REGION Network 32: "MFC-4024-T_DB"
   RUNG wire#powerrail
      "MFC-4024-T_DB"(Mode := 2, RAIVI :=, RAIVR :=, EnableHighAlarms :=, EnableLowAlarms :=, "TI Fail" :=, SAI =>)
   END_RUNG
   RUNG wire#powerrail
      I_Contact( false )
      { S7_GenerateENO := "TRUE" } Move(in := "MFC-4024_MB_R_DB".MB_Data.Buffer[2], out1 => "MFC-4024-T_DB".RAIVR)
   END_RUNG
   // the same network as SCL:
   "MFC-4024-T_DB"(Mode := 2);   // "TX-AI"
   IF NOT false THEN "MFC-4024-T_DB".RAIVR := "MFC-4024_MB_R_DB".MB_Data.Buffer[2]; END_IF;
END_REGION

REGION Network 33: "MFC-4025-T_DB"
   RUNG wire#powerrail
      "MFC-4025-T_DB"(Mode := 2, RAIVI :=, RAIVR :=, EnableHighAlarms :=, EnableLowAlarms :=, "TI Fail" :=, SAI =>)
   END_RUNG
   RUNG wire#powerrail
      I_Contact( false )
      { S7_GenerateENO := "TRUE" } Move(in := "MFC-4025_MB_R_DB".MB_Data.Buffer[2], out1 => "MFC-4025-T_DB".RAIVR)
   END_RUNG
   // the same network as SCL:
   "MFC-4025-T_DB"(Mode := 2);   // "TX-AI"
   IF NOT false THEN "MFC-4025-T_DB".RAIVR := "MFC-4025_MB_R_DB".MB_Data.Buffer[2]; END_IF;
END_REGION
END_FUNCTION

// folder: Analogs inputs/Trasmitters/VFD_Feedback Trasmitters

FUNCTION "VFDFeedbackTrasmitters" : Void   // FC14, LAD
TITLE = VFD Feedback
{ S7_Optimized_Access := 'TRUE' }
VERSION : 0.1
// Updated Date:
// Note:
   VAR_TEMP
      Alarms : Struct
         "T-101_AlarmsEnab" : Bool;
         "T-102_AlarmsEnab" : Bool;
         "R-201_AlarmsEnab" : Bool;
         "R-202_AlarmsEnab" : Bool;
         Centrifuge_AlarmsEnab : Bool;
      END_STRUCT;
      temporalvar : Int;
   END_VAR
BEGIN

REGION Network 1: Enable T-101 Agitator Alarms
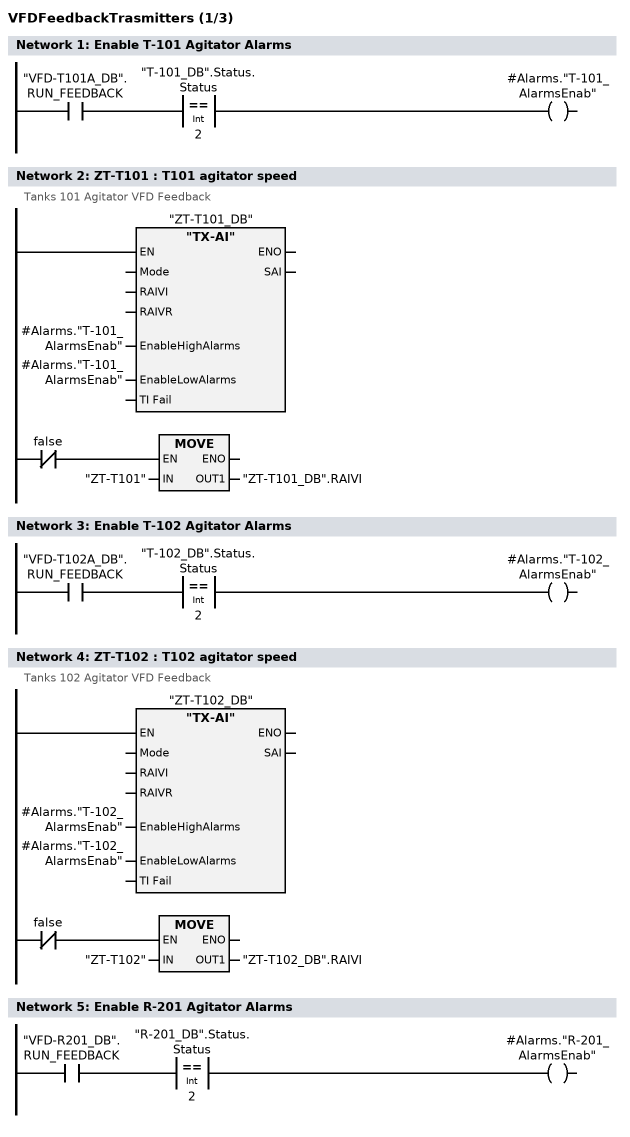
   RUNG wire#powerrail
      Contact( "VFD-T101A_DB".RUN_FEEDBACK )
      { S7_Templates := "SrcType := Int" } EQ_Contact(in1 := "T-101_DB".Status.Status, in2 := 2)
      Coil( #Alarms."T-101_AlarmsEnab" )
   END_RUNG
   // the same network as SCL:
   #Alarms."T-101_AlarmsEnab" := "VFD-T101A_DB".RUN_FEEDBACK AND ("T-101_DB".Status.Status = 2);
END_REGION

REGION Network 2: ZT-T101 : T101 agitator speed
   // Tanks 101 Agitator VFD Feedback
   RUNG wire#powerrail
      "ZT-T101_DB"(Mode :=, RAIVI :=, RAIVR :=, EnableHighAlarms := #Alarms."T-101_AlarmsEnab", EnableLowAlarms := #Alarms."T-101_AlarmsEnab", "TI Fail" :=, SAI =>)
   END_RUNG
   RUNG wire#powerrail
      I_Contact( false )
      { S7_GenerateENO := "TRUE" } Move(in := "ZT-T101", out1 => "ZT-T101_DB".RAIVI)
   END_RUNG
   // the same network as SCL:
   "ZT-T101_DB"(EnableHighAlarms := #Alarms."T-101_AlarmsEnab", EnableLowAlarms := #Alarms."T-101_AlarmsEnab");   // "TX-AI"
   IF NOT false THEN "ZT-T101_DB".RAIVI := "ZT-T101"; END_IF;
END_REGION

REGION Network 3: Enable T-102 Agitator Alarms
   RUNG wire#powerrail
      Contact( "VFD-T102A_DB".RUN_FEEDBACK )
      { S7_Templates := "SrcType := Int" } EQ_Contact(in1 := "T-102_DB".Status.Status, in2 := 2)
      Coil( #Alarms."T-102_AlarmsEnab" )
   END_RUNG
   // the same network as SCL:
   #Alarms."T-102_AlarmsEnab" := "VFD-T102A_DB".RUN_FEEDBACK AND ("T-102_DB".Status.Status = 2);
END_REGION

REGION Network 4: ZT-T102 : T102 agitator speed
   // Tanks 102 Agitator VFD Feedback
   RUNG wire#powerrail
      "ZT-T102_DB"(Mode :=, RAIVI :=, RAIVR :=, EnableHighAlarms := #Alarms."T-102_AlarmsEnab", EnableLowAlarms := #Alarms."T-102_AlarmsEnab", "TI Fail" :=, SAI =>)
   END_RUNG
   RUNG wire#powerrail
      I_Contact( false )
      { S7_GenerateENO := "TRUE" } Move(in := "ZT-T102", out1 => "ZT-T102_DB".RAIVI)
   END_RUNG
   // the same network as SCL:
   "ZT-T102_DB"(EnableHighAlarms := #Alarms."T-102_AlarmsEnab", EnableLowAlarms := #Alarms."T-102_AlarmsEnab");   // "TX-AI"
   IF NOT false THEN "ZT-T102_DB".RAIVI := "ZT-T102"; END_IF;
END_REGION

REGION Network 5: Enable R-201 Agitator Alarms
   RUNG wire#powerrail
      Contact( "VFD-R201_DB".RUN_FEEDBACK )
      { S7_Templates := "SrcType := Int" } EQ_Contact(in1 := "R-201_DB".Status.Status, in2 := 2)
      Coil( #Alarms."R-201_AlarmsEnab" )
   END_RUNG
   // the same network as SCL:
   #Alarms."R-201_AlarmsEnab" := "VFD-R201_DB".RUN_FEEDBACK AND ("R-201_DB".Status.Status = 2);
END_REGION

REGION Network 6: ZT-R201 : R201 agitator speed
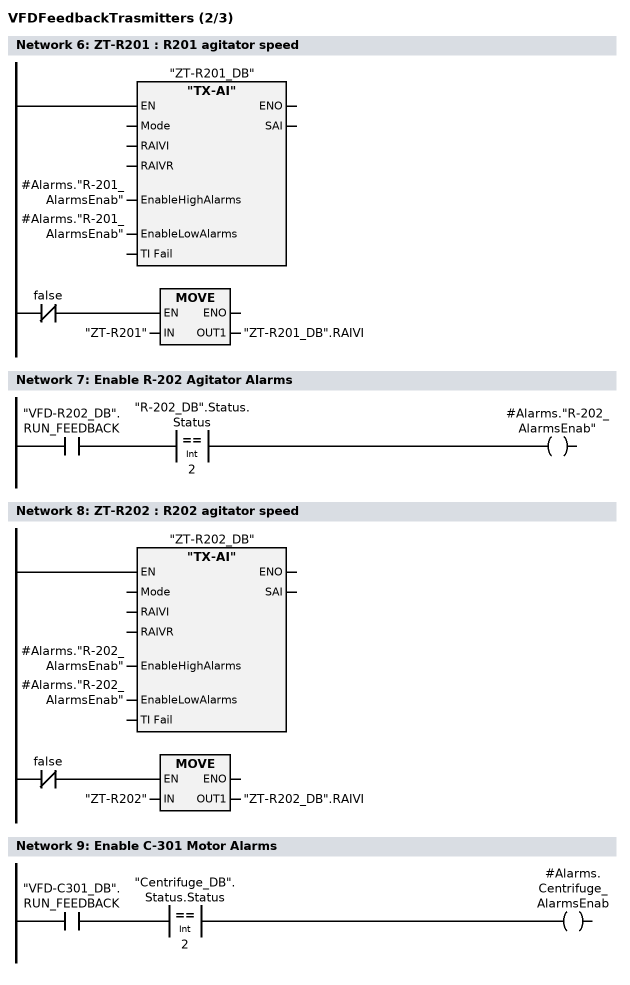
   RUNG wire#powerrail
      "ZT-R201_DB"(Mode :=, RAIVI :=, RAIVR :=, EnableHighAlarms := #Alarms."R-201_AlarmsEnab", EnableLowAlarms := #Alarms."R-201_AlarmsEnab", "TI Fail" :=, SAI =>)
   END_RUNG
   RUNG wire#powerrail
      I_Contact( false )
      { S7_GenerateENO := "TRUE" } Move(in := "ZT-R201", out1 => "ZT-R201_DB".RAIVI)
   END_RUNG
   // the same network as SCL:
   "ZT-R201_DB"(EnableHighAlarms := #Alarms."R-201_AlarmsEnab", EnableLowAlarms := #Alarms."R-201_AlarmsEnab");   // "TX-AI"
   IF NOT false THEN "ZT-R201_DB".RAIVI := "ZT-R201"; END_IF;
END_REGION

REGION Network 7: Enable R-202 Agitator Alarms
   RUNG wire#powerrail
      Contact( "VFD-R202_DB".RUN_FEEDBACK )
      { S7_Templates := "SrcType := Int" } EQ_Contact(in1 := "R-202_DB".Status.Status, in2 := 2)
      Coil( #Alarms."R-202_AlarmsEnab" )
   END_RUNG
   // the same network as SCL:
   #Alarms."R-202_AlarmsEnab" := "VFD-R202_DB".RUN_FEEDBACK AND ("R-202_DB".Status.Status = 2);
END_REGION

REGION Network 8: ZT-R202 : R202 agitator speed
   RUNG wire#powerrail
      "ZT-R202_DB"(Mode :=, RAIVI :=, RAIVR :=, EnableHighAlarms := #Alarms."R-202_AlarmsEnab", EnableLowAlarms := #Alarms."R-202_AlarmsEnab", "TI Fail" :=, SAI =>)
   END_RUNG
   RUNG wire#powerrail
      I_Contact( false )
      { S7_GenerateENO := "TRUE" } Move(in := "ZT-R202", out1 => "ZT-R202_DB".RAIVI)
   END_RUNG
   // the same network as SCL:
   "ZT-R202_DB"(EnableHighAlarms := #Alarms."R-202_AlarmsEnab", EnableLowAlarms := #Alarms."R-202_AlarmsEnab");   // "TX-AI"
   IF NOT false THEN "ZT-R202_DB".RAIVI := "ZT-R202"; END_IF;
END_REGION

REGION Network 9: Enable C-301 Motor Alarms
   RUNG wire#powerrail
      Contact( "VFD-C301_DB".RUN_FEEDBACK )
      { S7_Templates := "SrcType := Int" } EQ_Contact(in1 := "Centrifuge_DB".Status.Status, in2 := 2)
      Coil( #Alarms.Centrifuge_AlarmsEnab )
   END_RUNG
   // the same network as SCL:
   #Alarms.Centrifuge_AlarmsEnab := "VFD-C301_DB".RUN_FEEDBACK AND ("Centrifuge_DB".Status.Status = 2);
END_REGION

REGION Network 10: ZT-C-301 : C-301 Motorspeed
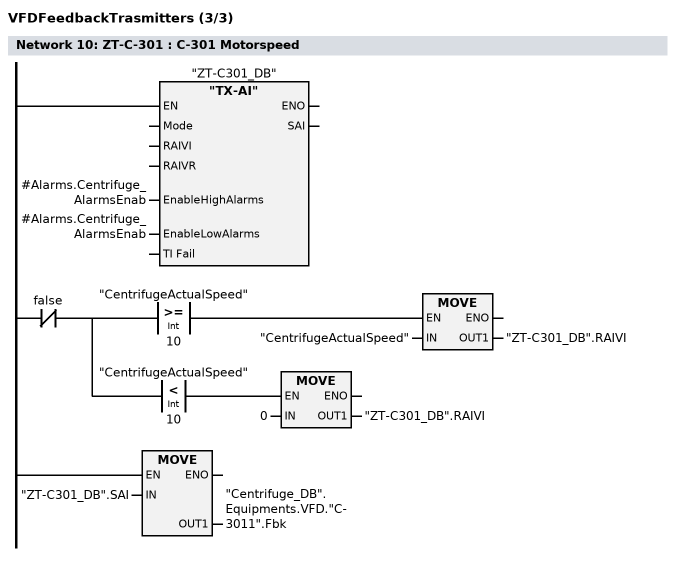
   RUNG wire#powerrail
      "ZT-C301_DB"(Mode :=, RAIVI :=, RAIVR :=, EnableHighAlarms := #Alarms.Centrifuge_AlarmsEnab, EnableLowAlarms := #Alarms.Centrifuge_AlarmsEnab, "TI Fail" :=, SAI =>)
   END_RUNG
   RUNG wire#powerrail
      I_Contact( false )
      wire#w1
      { S7_Templates := "SrcType := Int" } GE_Contact(in1 := "CentrifugeActualSpeed", in2 := 10)
      { S7_GenerateENO := "TRUE" } Move(in := "CentrifugeActualSpeed", out1 => "ZT-C301_DB".RAIVI)
   END_RUNG
   RUNG wire#w1
      { S7_Templates := "SrcType := Int" } LT_Contact(in1 := "CentrifugeActualSpeed", in2 := 10)
      { S7_GenerateENO := "TRUE" } Move(in := 0, out1 => "ZT-C301_DB".RAIVI)
   END_RUNG
   RUNG wire#powerrail
      Move(in := "ZT-C301_DB".SAI, out1 => "Centrifuge_DB".Equipments.VFD."C-3011".Fbk)
   END_RUNG
   // the same network as SCL:
   "ZT-C301_DB"(EnableHighAlarms := #Alarms.Centrifuge_AlarmsEnab,   // "TX-AI"
                EnableLowAlarms := #Alarms.Centrifuge_AlarmsEnab);
   IF NOT false AND ("CentrifugeActualSpeed" >= 10) THEN
       "ZT-C301_DB".RAIVI := "CentrifugeActualSpeed";
   END_IF;
   IF NOT false AND ("CentrifugeActualSpeed" < 10) THEN "ZT-C301_DB".RAIVI := 0; END_IF;
   "Centrifuge_DB".Equipments.VFD."C-3011".Fbk := "ZT-C301_DB".SAI;
END_REGION
END_FUNCTION

// folder: Analogs inputs/Trasmitters/Vibration Transmitter

FUNCTION "VibrationTransmitter" : Void   // FC107, LAD
{ S7_Optimized_Access := 'TRUE' }
VERSION : 0.1
BEGIN

REGION Network 1: Centrifuge Vibration Transmitter
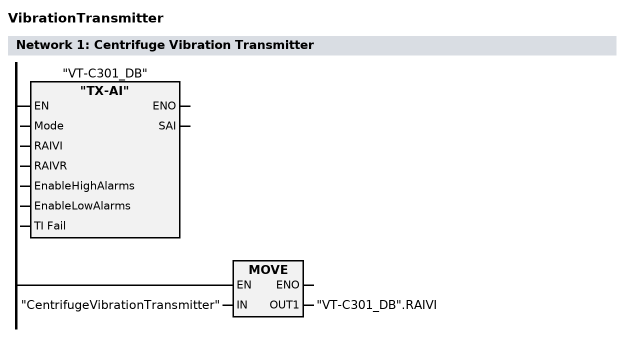
   RUNG wire#powerrail
      "VT-C301_DB"(Mode :=, RAIVI :=, RAIVR :=, EnableHighAlarms :=, EnableLowAlarms :=, "TI Fail" :=, SAI =>)
   END_RUNG
   RUNG wire#powerrail
      Move(in := "CentrifugeVibrationTransmitter", out1 => "VT-C301_DB".RAIVI)
   END_RUNG
   // the same network as SCL:
   "VT-C301_DB"();   // "TX-AI"
   "VT-C301_DB".RAIVI := "CentrifugeVibrationTransmitter";
END_REGION
END_FUNCTION

// folder: Calculations

FUNCTION_BLOCK "Array_Intergration"   // FB21, LAD
TITLE = Level to VFD Table
{ S7_Optimized_Access := 'TRUE' }
VERSION : 0.1
// Level to V FD Interpolation Table
   VAR_INPUT
      PV : Real;
      Ramp_UP : Bool := True;   // Ramp Up Sequence Enable
      Ramp_Down : Bool;   // Ramp Down Sequence Enable
   END_VAR
   VAR_OUTPUT
      SP : Real;
   END_VAR
   VAR
      FirstScan : Bool := TRUE;
      Number : UInt;
      "Array" : Array[0..#Array_Size] of Struct
         X : Real;   // Set Point for Level
         Y : Real;   // Output to Drive VFD
         X1 : Real;
         X2 : Real;
         Y1 : Real;
      END_STRUCT;
      TP_Up : IEC_TIMER;
      TP_Down : IEC_TIMER;
      Deadband : Struct
         UDW : Real := 0.5;   // Upper Deadband Width
         LDW : Real := 0.5;   // Lower Deadband Width
      END_STRUCT;
   END_VAR
   VAR_TEMP
      Trigger : Array[0..1] of Bool;
      Deadband_SP : Struct
         UDW : Real;   // Upper Deadband Width
         LDW : Real;   // Lower Deadband Width
      END_STRUCT;
      temp_CAl : Array[0..#Temp_Count] of Real;
   END_VAR
   VAR CONSTANT
      Array_Size : UInt := 4;
      TRigger_Count : UInt := 2;
      Temp_Count : UInt := 4;
   END_VAR
   VAR_TEMP   // added for the SCL form of the ladder/FBD networks
      _w1 : Bool;
      _w2 : Bool;
   END_VAR
   // "Array"[1].X := 20.0;
   // "Array"[2].X := 30.0;
   // "Array"[3].X := 40.0;
   // "Array"[4].X := 50.0;
   // TP_Up.PT := T#1ms;
   // TP_Down.PT := T#500ms;
BEGIN

REGION Network 1: First Scan
   // First Scan  Set array to Begining of the Table
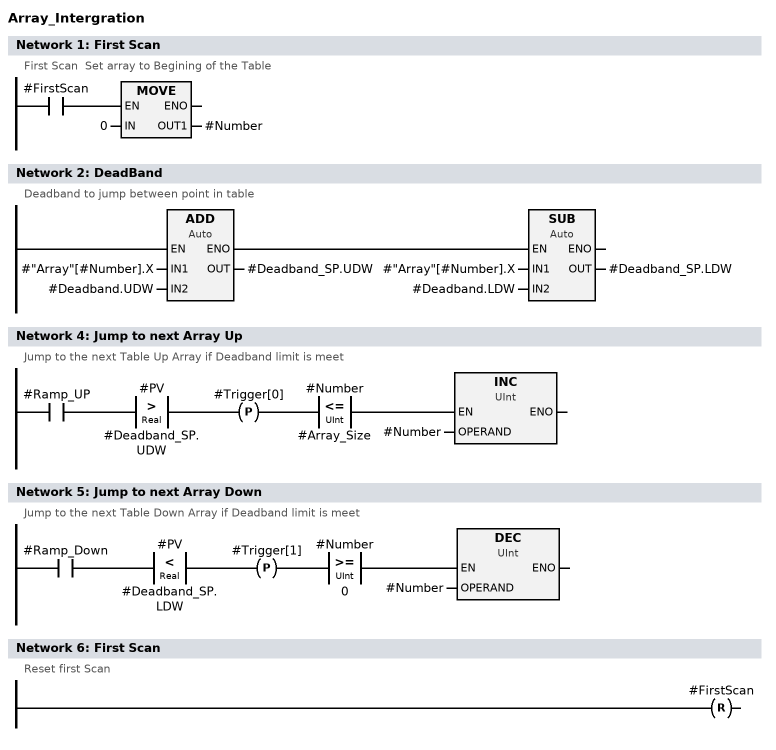
   RUNG wire#powerrail
      Contact( #FirstScan )
      { S7_GenerateENO := "TRUE" } Move(in := 0, out1 => #Number)
   END_RUNG
   // the same network as SCL:
   IF #FirstScan THEN #Number := 0; END_IF;
END_REGION

REGION Network 2: DeadBand
   // Deadband to jump between point in table
   RUNG wire#powerrail
      { S7_GenerateENO := "TRUE" } Add(in1 := #"Array"[#Number].X, in2 := #Deadband.UDW, out => #Deadband_SP.UDW)
      { S7_GenerateENO := "TRUE" } Sub(in1 := #"Array"[#Number].X, in2 := #Deadband.LDW, out => #Deadband_SP.LDW)
   END_RUNG
   // the same network as SCL:
   // ENO of a box is taken as its EN; it also drops when the box reports an error
   #Deadband_SP.UDW := #"Array"[#Number].X + #Deadband.UDW;
   #Deadband_SP.LDW := #"Array"[#Number].X - #Deadband.LDW;
END_REGION

REGION Network 3 (SCL): Table Calculation
   // Interpolation Formula implementation if the Ramp sequence is on and Deadband
   IF #Ramp_UP=TRUE AND #PV<=#Deadband_SP.UDW THEN
       // Interpolation Formula
       // Y = Y1 + (Y2 – Y1)/(X2 – X1) * (X * X1)
       #temp_CAl[0] := #Array[#Number].X * #Array[#Number].X1;// (X * X1)
       #temp_CAl[1] := #Array[#Number].X2 * #Array[#Number].X1;// (X2 – X1)
       #temp_CAl[2] := #Array[#Number].X2 * #Array[#Number].X1;// (Y2 – Y1)
       #temp_CAl[3] := #temp_CAl[1] / #temp_CAl[2];//(Y2 – Y1)/(X2 – X1)
       #temp_CAl[4] := #temp_CAl[3] * #temp_CAl[0];
       #SP := #Array[#Number].Y1 + #temp_CAl[4]; //SUM
   END_IF;
   IF #Ramp_Down=TRUE AND #PV>=#Deadband_SP.LDW THEN
       // Interpolation Formula
       // Y = Y1 + (Y2 – Y1)/(X2 – X1) * (X * X1)
       #temp_CAl[0] := #Array[#Number].X * #Array[#Number].X1;// (X * X1)
       #temp_CAl[1] := #Array[#Number].X2 * #Array[#Number].X1;// (X2 – X1)
       #temp_CAl[2] := #Array[#Number].X2 * #Array[#Number].X1;// (Y2 – Y1)
       #temp_CAl[3] := #temp_CAl[1] / #temp_CAl[2];//(Y2 – Y1)/(X2 – X1)
       #temp_CAl[4] := #temp_CAl[3] * #temp_CAl[0];
       #SP := #Array[#Number].Y1 + #temp_CAl[4]; //SUM
   END_IF;
END_REGION

REGION Network 4: Jump to next Array Up
   // Jump to the next Table Up Array if Deadband limit is meet
   RUNG wire#powerrail
      Contact( #Ramp_UP )
      { S7_Templates := "SrcType := Real" } GT_Contact(in1 := #PV, in2 := #Deadband_SP.UDW)
      P_Trig( #Trigger[0] )
      { S7_Templates := "SrcType := UInt" } LE_Contact(in1 := #Number, in2 := #Array_Size)
      { S7_Templates := "DestType := UInt"; S7_GenerateENO := "TRUE" } Inc( #Number )
   END_RUNG
   // the same network as SCL:
   #_w1 := #Ramp_UP AND (#PV > #Deadband_SP.UDW);
   #_w2 := #_w1 AND NOT #Trigger[0];   // rising edge
   #Trigger[0] := #_w1;
   IF #_w2 AND (#Number <= #Array_Size) THEN #Number := #Number + 1; END_IF;
END_REGION

REGION Network 5: Jump to next Array Down
   // Jump to the next Table Down Array if Deadband limit is meet
   RUNG wire#powerrail
      Contact( #Ramp_Down )
      { S7_Templates := "SrcType := Real" } LT_Contact(in1 := #PV, in2 := #Deadband_SP.LDW)
      P_Trig( #Trigger[1] )
      { S7_Templates := "SrcType := UInt" } GE_Contact(in1 := #Number, in2 := 0)
      { S7_Templates := "DestType := UInt"; S7_GenerateENO := "TRUE" } Dec( #Number )
   END_RUNG
   // the same network as SCL:
   #_w1 := #Ramp_Down AND (#PV < #Deadband_SP.LDW);
   #_w2 := #_w1 AND NOT #Trigger[1];   // rising edge
   #Trigger[1] := #_w1;
   IF #_w2 AND (#Number >= 0) THEN #Number := #Number - 1; END_IF;
END_REGION

REGION Network 6: First Scan
   // Reset first Scan
   RUNG wire#powerrail
      R_Coil( #FirstScan )
   END_RUNG
   // the same network as SCL:
   #FirstScan := FALSE;
END_REGION
END_FUNCTION_BLOCK

FUNCTION_BLOCK "Tank_Calculation_FB"   // FB22, LAD
{ S7_Optimized_Access := 'TRUE' }
VERSION : 0.1
   VAR_INPUT
      Mode : UInt;   // Type of Tank mode: 1= Vertical Capsule Tank
      Level : Real;
   END_VAR
   VAR_OUTPUT
      ScaleVolume : Real;
   END_VAR
   VAR
      "Vertical Capsule Tank" : Struct
         Enable : Bool;
         "case" : USInt;   // Mode: | Vcylpartial=1 | Vcylpartial & Vbottom_head_partial = 2 | Vcylpartial & Vtop_head_partial = 3 | Vcyl_total = 4 |
         Static_1 : USInt;   // tank internal diameter
         DiameterCylindrical : UInt;
         Height : UInt;
      END_STRUCT;
   END_VAR
   VAR_TEMP
      "Case" : USInt;
      Vcylpartial : Real;
      TEmp : Real;
      temp_CAl : Array[0..#Temp_Count] of Real;
   END_VAR
   VAR CONSTANT
      "Vertical Capsule Tank_1" : UInt := 1;
      MAthPi : Real := 3.14;
      Temp_Count : UInt := 4;
   END_VAR
BEGIN

REGION Network 1: Mode1: Selected
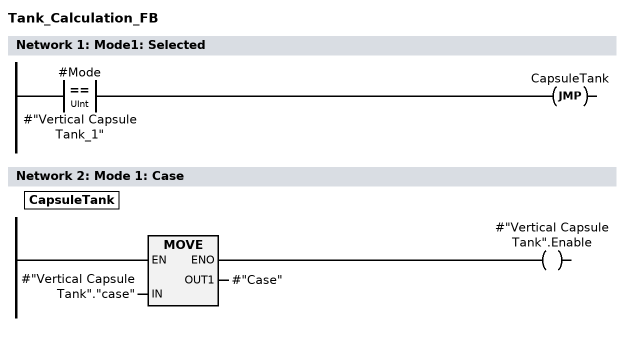
   RUNG wire#powerrail
      { S7_Templates := "SrcType := UInt" } EQ_Contact(in1 := #Mode, in2 := #"Vertical Capsule Tank_1")
      JumpCoil( CapsuleTank )
   END_RUNG
   // the same network as SCL:
   IF #Mode = #"Vertical Capsule Tank_1" THEN GOTO CapsuleTank; END_IF;
END_REGION

REGION Network 2: Mode 1: Case
   Label( CapsuleTank )
   RUNG wire#powerrail
      { S7_GenerateENO := "TRUE" } Move(in := #"Vertical Capsule Tank"."case", out1 => #"Case")
      Coil( #"Vertical Capsule Tank".Enable )
   END_RUNG
   // the same network as SCL:
   // ENO of a box is taken as its EN; it also drops when the box reports an error
   CapsuleTank:
   #"Case" := #"Vertical Capsule Tank"."case";
   #"Vertical Capsule Tank".Enable := TRUE;
END_REGION

REGION Network 3 (SCL): Vertical Capsule Tank CAlculation
   CASE #Case OF
       1:(*Mode:Partial Volume horizontal Cylinderical Calculation
       Note: Calculation For the cylindrical part Of the tank only 
             does not Contain Top Head or Botton Head of vessel
       Formula: Vcylpartial=π*〖ID〗^2/4*Lv*)
           #temp_CAl[0] := #"Vertical Capsule Tank".DiameterCylindrical / 2;//Radius /cylindrical
           #temp_CAl[1] := #MAthPi * #temp_CAl[0] ** 2 * (#Level - 2 * #temp_CAl[0]);// Volume Cylinderical  
           #temp_CAl[2] := #Level/ (#MAthPi * #temp_CAl[0] ** 2);// Liquid Level
           #Vcylpartial := #Level - (#temp_CAl[2]);// Current Level
           #ScaleVolume := #Vcylpartial;// Move To Volume
           ;
       2:  (*Mode: The liquid level is in the Botton head of the vessel to the top of the Cylinderical part of the Vessel the top head of the Vessel not  *)
           IF #Level >= 0 AND #Level <= 20 THEN
               // From 0 to 20 The liquid level is low, within the bottom head of the vessel
             //  #temp_CAl[0] := #MAthPi/6*(3*)  ;
             //  #Vbottom_head = 
               ;
           ELSE

               ;
           END_IF;


           ;
       3:  // The liquid level is reaching the top head of the vessel
           ;
       ELSE  // Set Case Value to 0
           #Case := 0;
           ;
   END_CASE;
END_REGION
END_FUNCTION_BLOCK

FUNCTION_BLOCK "Array_Intergration_B"   // FB23, LAD
TITLE = Level to VFD Table
{ S7_Optimized_Access := 'TRUE' }
VERSION : 0.1
// Level to V FD Interpolation Table
   VAR_INPUT
      PV : Int;
      Ramp_UP : Bool := True;   // Ramp Up Sequence Enable
      Ramp_Down : Bool;   // Ramp Down Sequence Enable
   END_VAR
   VAR_OUTPUT
      SP : Real;
   END_VAR
   VAR
      FirstScan : Bool := TRUE;
      Number : UInt;
      "X Axis Max" : Int := 100;
      "Y Axis max" : Int := 4000;
      "array of X" : Array[0..#Array_Size] of Int;   // Level Setpoints
      "array of Y" : Array[0..#Array_Size] of Int;   // RPM Sepoints
      "Array" : Array[0..#Array_Size] of Struct
         X : Int;   // Set Point for Level
         Y : Int;   // Output to Drive VFD
         X1 : Int;
         X2 : Int;
         Y1 : Int;
         Y2 : Int;
      END_STRUCT;
      Formula : Struct
         X : Int;   // Set Point for Level
         Y : Int;   // Output to Drive VFD
         X1 : Int;
         X2 : Int;
         Y1 : Int;
         Y2 : Int;
      END_STRUCT;
      TP_Up : IEC_TIMER;
      TP_Down : IEC_TIMER;
      Deadband : Struct
         UDW : Real := 0.5;   // Upper Deadband Width
         LDW : Real := 0.5;   // Lower Deadband Width
      END_STRUCT;
   END_VAR
   VAR_TEMP
      Trigger : Array[0..1] of Bool;
      Deadband_SP : Struct
         UDW : Real;   // Upper Deadband Width
         LDW : Real;   // Lower Deadband Width
      END_STRUCT;
      temp_CAl : Array[0..#Temp_Count] of Real;
   END_VAR
   VAR CONSTANT
      Array_Size : UInt := 4;
      TRigger_Count : UInt := 2;
      Temp_Count : UInt := 5;
      RMP : UInt := 3000;
   END_VAR
   // TP_Up.PT := T#1ms;
   // TP_Down.PT := T#500ms;
   // "array of X"[0] := 20;
   // "array of X"[1] := 30;
   // "array of X"[2] := 40;
   // "array of X"[3] := 50;
   // "array of X"[4] := 60;
   // "array of Y"[0] := 500;
   // "array of Y"[1] := 1000;
   // "array of Y"[2] := 1500;
   // "array of Y"[3] := 2000;
   // "array of Y"[4] := 1500;
BEGIN

REGION Network 1: First Scan
   // First Scan  Set array to Begining of the Table
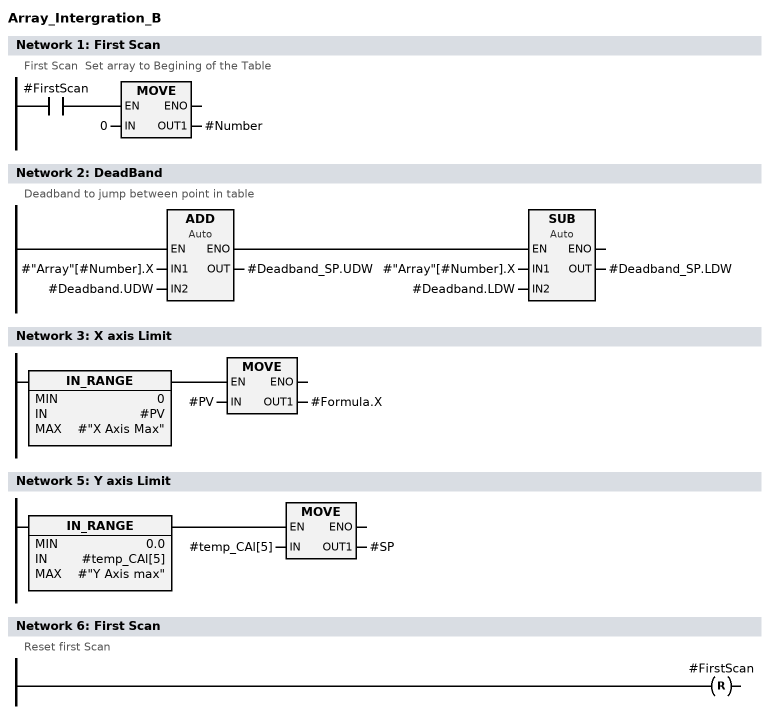
   RUNG wire#powerrail
      Contact( #FirstScan )
      { S7_GenerateENO := "TRUE" } Move(in := 0, out1 => #Number)
   END_RUNG
   // the same network as SCL:
   IF #FirstScan THEN #Number := 0; END_IF;
END_REGION

REGION Network 2: DeadBand
   // Deadband to jump between point in table
   RUNG wire#powerrail
      { S7_GenerateENO := "TRUE" } Add(in1 := #"Array"[#Number].X, in2 := #Deadband.UDW, out => #Deadband_SP.UDW)
      { S7_GenerateENO := "TRUE" } Sub(in1 := #"Array"[#Number].X, in2 := #Deadband.LDW, out => #Deadband_SP.LDW)
   END_RUNG
   // the same network as SCL:
   // ENO of a box is taken as its EN; it also drops when the box reports an error
   #Deadband_SP.UDW := #"Array"[#Number].X + #Deadband.UDW;
   #Deadband_SP.LDW := #"Array"[#Number].X - #Deadband.LDW;
END_REGION

REGION Network 3: X axis Limit
   RUNG wire#powerrail
      { S7_Templates := "SrcType := Int" } InRange(min := 0, in := #PV, max := #"X Axis Max")
      { S7_GenerateENO := "TRUE" } Move(in := #PV, out1 => #Formula.X)
   END_RUNG
   // the same network as SCL:
   IF (0 <= #PV) AND (#PV <= #"X Axis Max") THEN #Formula.X := #PV; END_IF;
END_REGION

REGION Network 4 (SCL): Table Calculation
   // Interpolation Formula implementation if the Ramp sequence is on and Deadband
   // Interpolation Formula
   // Y = Y1 + (Y2 – Y1)/(X2 – X1) * (X * X1)
   #Formula.Y1 := #"array of Y"[0];
   #Formula.X1 := #"array of X"[0];
   #Formula.Y2 := #"array of Y"[1];
   #Formula.X2 := #"array of X"[1];
   #temp_CAl[0] := #Formula.Y2 * #Formula.Y1;// (Y2 – Y1)
   #temp_CAl[1] := #Formula.X2 - #Formula.X1;// (X2 – X1)
   #temp_CAl[2] := #Formula.X * #Formula.X1;// (X * X1)
   #temp_CAl[3] := #temp_CAl[0] / #temp_CAl[1];//(Y2 – Y1)/(X2 – X1)
   #temp_CAl[4] := #temp_CAl[3] * #temp_CAl[2];//(Y2 – Y1)/(X2 – X1) * (X * X1)
   #temp_CAl[5] := #Formula.Y1 + #temp_CAl[4];//Y1 + (Y2 – Y1)/(X2 – X1) * (X * X1)
END_REGION

REGION Network 5: Y axis Limit
   RUNG wire#powerrail
      { S7_Templates := "SrcType := Real" } InRange(min := 0.0, in := #temp_CAl[5], max := #"Y Axis max")
      { S7_GenerateENO := "TRUE" } Move(in := #temp_CAl[5], out1 => #SP)
   END_RUNG
   // the same network as SCL:
   IF (0.0 <= #temp_CAl[5]) AND (#temp_CAl[5] <= #"Y Axis max") THEN #SP := #temp_CAl[5]; END_IF;
END_REGION

REGION Network 6: First Scan
   // Reset first Scan
   RUNG wire#powerrail
      R_Coil( #FirstScan )
   END_RUNG
   // the same network as SCL:
   #FirstScan := FALSE;
END_REGION
END_FUNCTION_BLOCK

FUNCTION_BLOCK "Volume_Calculation"   // FB25, SCL
{ S7_Optimized_Access := 'TRUE' }
VERSION : 0.1
   VAR_INPUT
      Input : Int;
      Input_Max : Real;
      Input_Min : Real;
   END_VAR
   VAR_OUTPUT
      "Volume (L)" : Real;   // Valume in Gallons
      "Volume (Gal)" : Real;   // Volume in Liters
   END_VAR
   VAR
      CurrentCylinderVolume : Struct   // Actual Volumeof the Cylinder
         L : Real;
         Gal : Real;
      END_STRUCT;
      LevelInp : Int;
      Dumm : Word;
      Dumm2 : Word;
   END_VAR
   VAR CONSTANT
      aLiter_To_Gallon : Real := 0.264;   // 1 Liter is equal to 0.264 Gallons
      Pi : Real := 3.1416;
      aft_To_cm : Real := 30.48;
   END_VAR
BEGIN




   IF #Input >= 0 AND #Input <= 27648 THEN

       //#LevelInp := REAL_TO_INT(IN := #Level_inch);
       //#Dumm := SCALE(IN := #LevelInp, HI_LIM := #"HI_Vol (Gal)", LO_LIM := #"LO_Vol (Gal)", BIPOLAR := False, OUT => #"Volume (Gal)");
       #Dumm2 := SCALE(IN := #Input, HI_LIM := #Input_Max, LO_LIM := #Input_Min, BIPOLAR := FALSE, OUT => #CurrentCylinderVolume.L);




       #CurrentCylinderVolume.Gal := #CurrentCylinderVolume.L / 3.785; //To convert to Galons ;1 Gal = 3.785 Liters

       #"Volume (L)" := #CurrentCylinderVolume.L;
       #"Volume (Gal)" := #CurrentCylinderVolume.Gal;

   ELSE
       #"Volume (L)" := 0.0;
       #"Volume (Gal)" := 0.0;

   END_IF;
END_FUNCTION_BLOCK

FUNCTION_BLOCK "INTEGRATE_FB"   // FB26, SCL
{ S7_Optimized_Access := 'TRUE' }
VERSION : 0.1
   VAR_INPUT
      rYin : Real;   // Input Variable (e.g. flow)
      rTd : Real;   // Sampling time period [e.g. s]
      rYk : Real;   // Y factor (to convert Yin to a per-sampling-time rate) [e.g. Yunits/s]
      boEn : Bool;   // Enable integration function
      boRst : Bool;   // Reset integrated value
   END_VAR
   VAR_OUTPUT
      rYout : Real;   // Result of integrated function (= area below Yin) (result)
   END_VAR
   VAR
      rYs : Real;   // Result of integrated function (= area below Yin) (internal)
      TempVal : Real;   // Per-Sampling-Time Rate
   END_VAR
BEGIN
   (*
   This function implements an Integration Function.

   Function must be called from a time-interrupt OB

   Call Example:

         CALL  "INTEGRATE_FB" , "INTEGRATE_DB"
          diYin:="BXP_INTEGRATE_DB".diYin
          rTd  :=1.000000e-001             //  Sampling rate: 0.1 [s]
          rYk  :=2.777777e-004             //  1 [unit/h] = 1/3600
          boEn :="BXP_INTEGRATE_DB".boEn
          boRst:="BXP_INTEGRATE_DB".boRst
          diYs :="BXP_INTEGRATE_DB".diYs

   rTd:= Sampling rate: 0.1 [s]
   rYk:=   1 [l/h] = 1/3600 [l/s] or [l/m] *This value depend of the units from the Flow meter
   *)

   IF NOT #boRst THEN //Reset?
       IF #boEn THEN   //// Function Enabled?
           //Integrate
           #TempVal := #rYin * #rYk;   //Y factor (to convert Yin to a per-sampling-time rate) [e.g. Yunits/s]
           #TempVal := #TempVal * #rTd;

           #rYs := #rYs + #TempVal;    //Result of integrated function (= area below Yin) (internal)

           #rYout := #rYs;    //Result of integrated function (= area below Yin) (result)

       ELSE
           //// Return last computed value when function disabled
           #rYs := #rYs;
           #rYout := #rYs;
       END_IF;
   ELSE
       // Reset accumulated value when reset
       #rYs := 0.0;
       #rYout := #rYs;

   END_IF;
END_FUNCTION_BLOCK

FUNCTION "Tank_Calculation" : Void   // FC18, LAD
{ S7_Optimized_Access := 'TRUE' }
VERSION : 0.1
BEGIN

REGION Network 1 (SCL): LT-1011 : T-101 X Material Volume Calculation
END_REGION
END_FUNCTION

FUNCTION "Calculator_Caller" : Void   // FC103, LAD
{ S7_Optimized_Access := 'TRUE' }
VERSION : 0.1
BEGIN

REGION Network 1
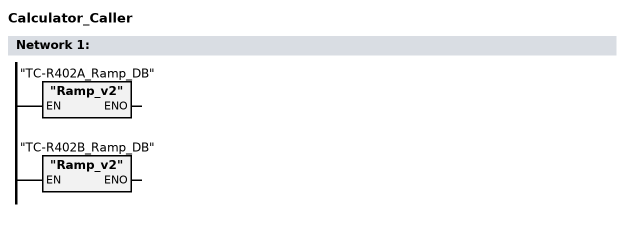
   RUNG wire#powerrail
      "TC-R402A_Ramp_DB"()
   END_RUNG
   RUNG wire#powerrail
      "TC-R402B_Ramp_DB"()
   END_RUNG
   // the same network as SCL:
   "TC-R402A_Ramp_DB"();   // "Ramp_v2"
   "TC-R402B_Ramp_DB"();   // "Ramp_v2"
END_REGION
END_FUNCTION

// folder: Cause&EffectMatrix

FUNCTION_BLOCK "CauseAndEffect"   // FB5, CEM
{ S7_Optimized_Access := 'TRUE' }
VERSION : 0.1
   VAR_INPUT
      C1 : Bool;
   END_VAR
   VAR_OUTPUT
      E1 : Bool;
   END_VAR
   VAR
      RTData : Struct
         CauseActive : Array[0..7] of Bool;
         CauseActiveCompressed : Array[0..0] of Byte;
         EffectActive : Array[0..7] of Bool;
         EffectActiveCompressed : Array[0..0] of Byte;
         Intersections : Array[0..5] of Byte;   // (start values stored as a binary block, not shown)
         History : Array[0..0] of Byte;
         RunFlag : Bool;
         "Timer" : IEC_TIMER;
         CycleStartTime : Time;
      END_STRUCT;
      Cause1 : CEM_Cause;
      Effect1 : CEM_Effect;
   END_VAR
BEGIN

REGION Network 1
   // network source EffectGroups not rendered
END_REGION

REGION Network 2
   // network source CauseGroups not rendered
END_REGION

REGION Network 3
   // network source Cause not rendered
END_REGION

REGION Network 4
   // network source Effect not rendered
END_REGION
END_FUNCTION_BLOCK

// folder: Diagnostic

FUNCTION_BLOCK "diag"   // FB14, LAD
{ S7_Optimized_Access := 'TRUE' }
VERSION : 0.1
   VAR
      SHUTDOWN : Bool;
      PS1 : Bool;
      PS2 : Bool;
   END_VAR
BEGIN

REGION Network 1: PWR SUPPLY SIGNAL
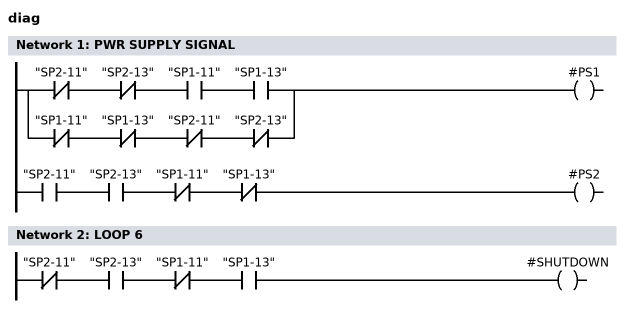
   RUNG wire#powerrail
      I_Contact( "SP2-11" )
      I_Contact( "SP2-13" )
      Contact( "SP1-11" )
      Contact( "SP1-13" )
      wire#w1
      Coil( #PS1 )
   END_RUNG
   RUNG wire#powerrail
      I_Contact( "SP1-11" )
      I_Contact( "SP1-13" )
      I_Contact( "SP2-11" )
      I_Contact( "SP2-13" )
   END_RUNG wire#w1
   RUNG wire#powerrail
      Contact( "SP2-11" )
      Contact( "SP2-13" )
      I_Contact( "SP1-11" )
      I_Contact( "SP1-13" )
      Coil( #PS2 )
   END_RUNG
   // the same network as SCL:
   #PS1 := (NOT "SP2-11" AND NOT "SP2-13" AND "SP1-11" AND "SP1-13") OR (NOT "SP1-11" AND NOT "SP1-13" AND NOT "SP2-11" AND NOT "SP2-13");
   #PS2 := "SP2-11" AND "SP2-13" AND NOT "SP1-11" AND NOT "SP1-13";
END_REGION

REGION Network 2: LOOP 6
   RUNG wire#powerrail
      I_Contact( "SP2-11" )
      Contact( "SP2-13" )
      I_Contact( "SP1-11" )
      Contact( "SP1-13" )
      Coil( #SHUTDOWN )
   END_RUNG
   // the same network as SCL:
   #SHUTDOWN := NOT "SP2-11" AND "SP2-13" AND NOT "SP1-11" AND "SP1-13";
END_REGION

REGION Network 3: LOOP 7
END_REGION
END_FUNCTION_BLOCK

// folder: ESD

FUNCTION "Interlocks_FB" : Void   // FC20, LAD
{ S7_Optimized_Access := 'TRUE' }
VERSION : 0.1
   VAR_TEMP
      REAL_1 : Real;
      INT_1 : Real;
      INT_2 : Real;
   END_VAR
BEGIN

REGION Network 1: T-101 Mix & Wash X material
   // loop 1 &2